REGION Network 6: GET NEXT STATION
   RUNG wire#powerrail
      P_Contact(operand := #settings.viewingStation.next.actuate, bit := #old.nextPress)
      wire#w1
      { S7_Templates := "SrcType := Int" } NE_Contact(in1 := #settings.stations.selCount, in2 := 0)
      "Get Station Selection Number"(next := TRUE, prev := FALSE, stations := #stations, selStnNumber := #settings.stations.selNumber)
   END_RUNG
   RUNG wire#powerrail
      { S7_Templates := "SrcType := Int" } NE_Contact(in1 := #settings.stations.selCount, in2 := #old.selStnCount)
   END_RUNG wire#w1
   // the same network as SCL:
   #_w1 := #settings.viewingStation.next.actuate AND NOT #old.nextPress;   // rising edge of #settings.viewingStation.next.actuate
   #old.nextPress := #settings.viewingStation.next.actuate;
   IF (#_w1 OR (#settings.stations.selCount <> #old.selStnCount)) AND (#settings.stations.selCount <> 0) THEN
       "Get Station Selection Number"(next := TRUE,
                               prev := FALSE,
                               stations := #stations,
                               selStnNumber := #settings.stations.selNumber);
   END_IF;
END_REGION

REGION Network 7: ANIMATE: NEXT STATION BUTTON
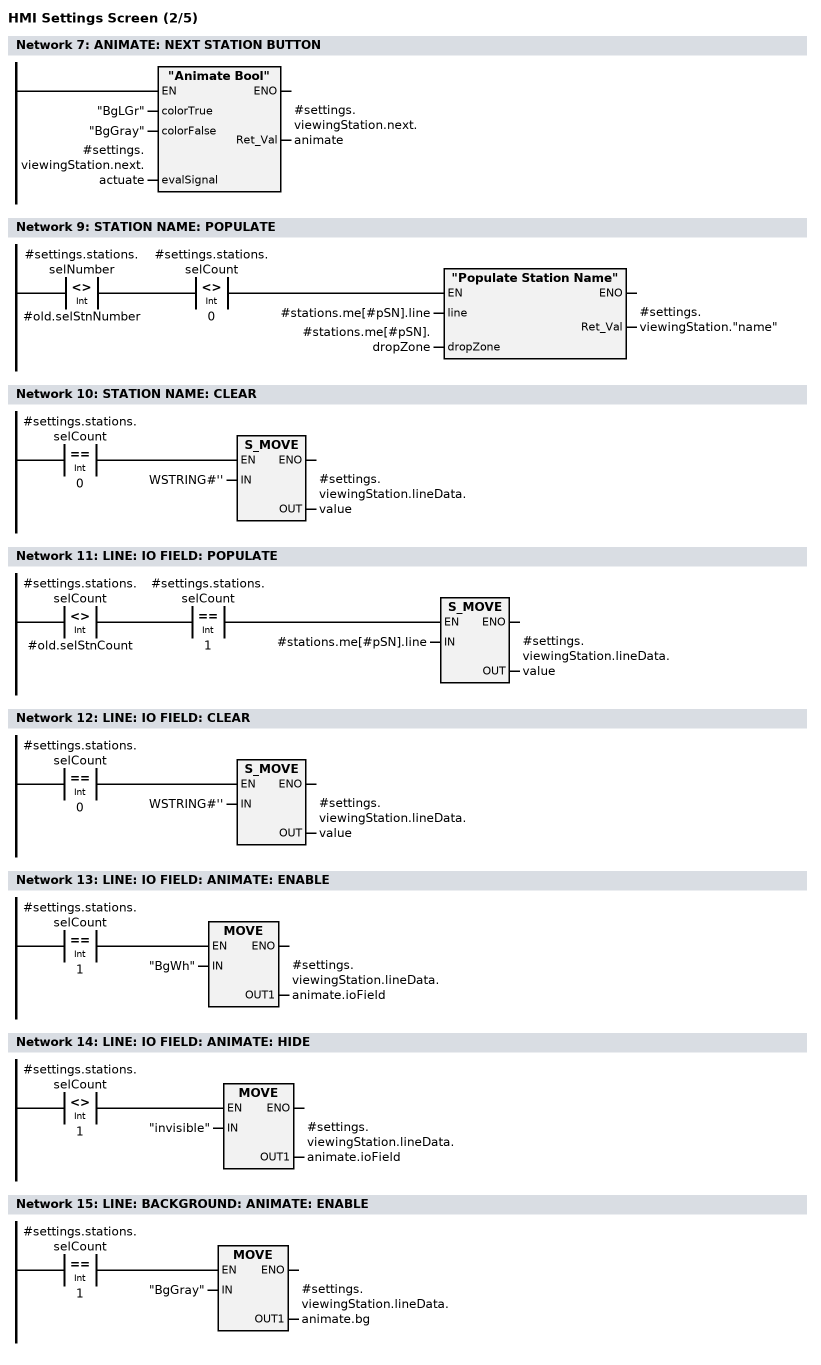
   RUNG wire#powerrail
      "Animate Bool"(colorTrue := "BgLGr", colorFalse := "BgGray", evalSignal := #settings.viewingStation.next.actuate, Ret_Val => #settings.viewingStation.next.animate)
   END_RUNG
   // the same network as SCL:
   #settings.viewingStation.next.animate := "Animate Bool"(colorTrue := "BgLGr",
                           colorFalse := "BgGray",
                           evalSignal := #settings.viewingStation.next.actuate);
END_REGION

REGION Network 8 (SCL): COPY TO POINTERS
   #pSN := #settings.stations.selNumber;
   #pBN := #settings.kp8.selBtnNumber;
END_REGION

REGION Network 9: STATION NAME: POPULATE
   RUNG wire#powerrail
      { S7_Templates := "SrcType := Int" } NE_Contact(in1 := #settings.stations.selNumber, in2 := #old.selStnNumber)
      { S7_Templates := "SrcType := Int" } NE_Contact(in1 := #settings.stations.selCount, in2 := 0)
      "Populate Station Name"(line := #stations.me[#pSN].line, dropZone := #stations.me[#pSN].dropZone, Ret_Val => #settings.viewingStation."name")
   END_RUNG
   // the same network as SCL:
   IF (#settings.stations.selNumber <> #old.selStnNumber) AND (#settings.stations.selCount <> 0) THEN
       #settings.viewingStation."name" := "Populate Station Name"(line := #stations.me[#pSN].line,
                               dropZone := #stations.me[#pSN].dropZone);
   END_IF;
END_REGION

REGION Network 10: STATION NAME: CLEAR
   RUNG wire#powerrail
      { S7_Templates := "SrcType := Int" } EQ_Contact(in1 := #settings.stations.selCount, in2 := 0)
      S_Move(in := WSTRING#'', out => #settings.viewingStation.lineData.value)
   END_RUNG
   // the same network as SCL:
   IF #settings.stations.selCount = 0 THEN #settings.viewingStation.lineData.value := WSTRING#''; END_IF;
END_REGION

REGION Network 11: LINE: IO FIELD: POPULATE
   RUNG wire#powerrail
      { S7_Templates := "SrcType := Int" } NE_Contact(in1 := #settings.stations.selCount, in2 := #old.selStnCount)
      { S7_Templates := "SrcType := Int" } EQ_Contact(in1 := #settings.stations.selCount, in2 := 1)
      S_Move(in := #stations.me[#pSN].line, out => #settings.viewingStation.lineData.value)
   END_RUNG
   // the same network as SCL:
   IF (#settings.stations.selCount <> #old.selStnCount) AND (#settings.stations.selCount = 1) THEN
       #settings.viewingStation.lineData.value := #stations.me[#pSN].line;
   END_IF;
END_REGION

REGION Network 12: LINE: IO FIELD: CLEAR
   RUNG wire#powerrail
      { S7_Templates := "SrcType := Int" } EQ_Contact(in1 := #settings.stations.selCount, in2 := 0)
      S_Move(in := WSTRING#'', out => #settings.viewingStation.lineData.value)
   END_RUNG
   // the same network as SCL:
   IF #settings.stations.selCount = 0 THEN #settings.viewingStation.lineData.value := WSTRING#''; END_IF;
END_REGION

REGION Network 13: LINE: IO FIELD: ANIMATE: ENABLE
   RUNG wire#powerrail
      { S7_Templates := "SrcType := Int" } EQ_Contact(in1 := #settings.stations.selCount, in2 := 1)
      Move(in := "BgWh", out1 => #settings.viewingStation.lineData.animate.ioField)
   END_RUNG
   // the same network as SCL:
   IF #settings.stations.selCount = 1 THEN
       #settings.viewingStation.lineData.animate.ioField := "BgWh";
   END_IF;
END_REGION

REGION Network 14: LINE: IO FIELD: ANIMATE: HIDE
   RUNG wire#powerrail
      { S7_Templates := "SrcType := Int" } NE_Contact(in1 := #settings.stations.selCount, in2 := 1)
      Move(in := "invisible", out1 => #settings.viewingStation.lineData.animate.ioField)
   END_RUNG
   // the same network as SCL:
   IF #settings.stations.selCount <> 1 THEN
       #settings.viewingStation.lineData.animate.ioField := "invisible";
   END_IF;
END_REGION

REGION Network 15: LINE: BACKGROUND: ANIMATE: ENABLE
   RUNG wire#powerrail
      { S7_Templates := "SrcType := Int" } EQ_Contact(in1 := #settings.stations.selCount, in2 := 1)
      Move(in := "BgGray", out1 => #settings.viewingStation.lineData.animate.bg)
   END_RUNG
   // the same network as SCL:
   IF #settings.stations.selCount = 1 THEN #settings.viewingStation.lineData.animate.bg := "BgGray"; END_IF;
END_REGION

REGION Network 16: LINE: BACKGROUND: ANIMATE: HIDE
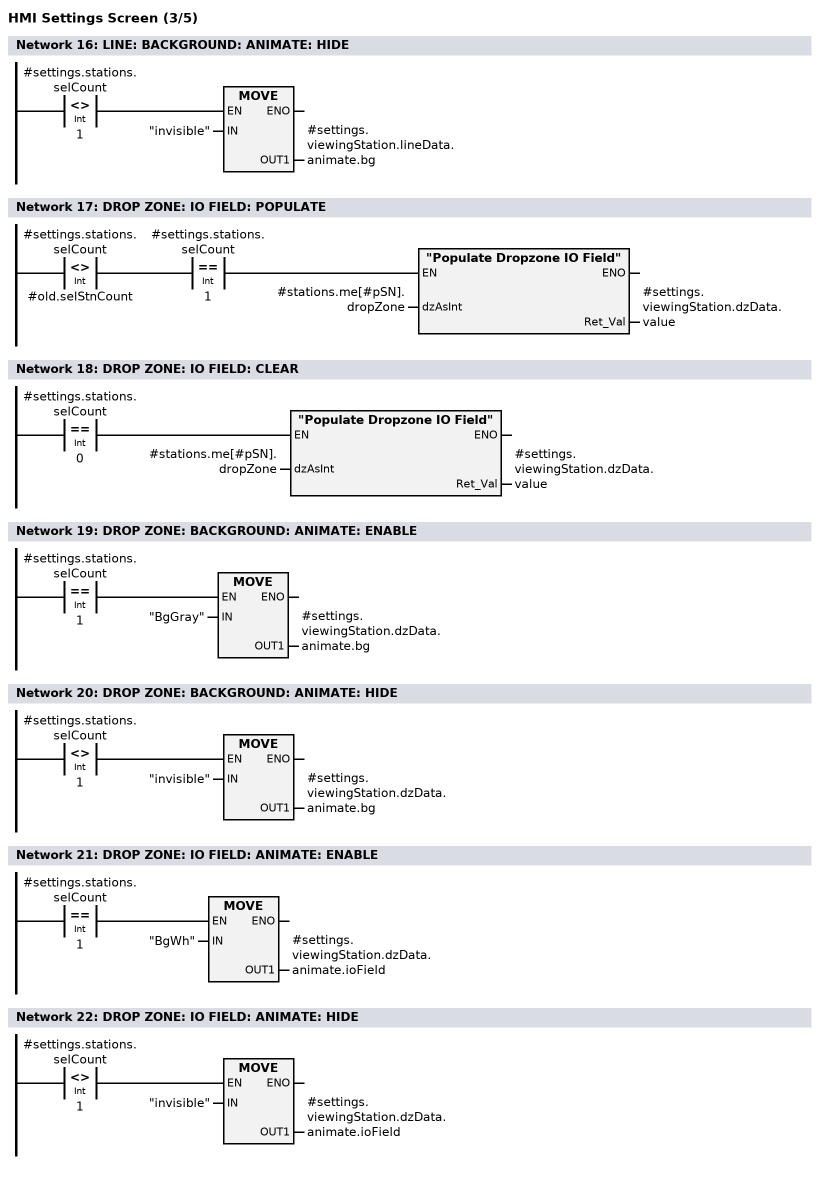
   RUNG wire#powerrail
      { S7_Templates := "SrcType := Int" } NE_Contact(in1 := #settings.stations.selCount, in2 := 1)
      Move(in := "invisible", out1 => #settings.viewingStation.lineData.animate.bg)
   END_RUNG
   // the same network as SCL:
   IF #settings.stations.selCount <> 1 THEN
       #settings.viewingStation.lineData.animate.bg := "invisible";
   END_IF;
END_REGION

REGION Network 17: DROP ZONE: IO FIELD: POPULATE
   RUNG wire#powerrail
      { S7_Templates := "SrcType := Int" } NE_Contact(in1 := #settings.stations.selCount, in2 := #old.selStnCount)
      { S7_Templates := "SrcType := Int" } EQ_Contact(in1 := #settings.stations.selCount, in2 := 1)
      "Populate Dropzone IO Field"(dzAsInt := #stations.me[#pSN].dropZone, Ret_Val => #settings.viewingStation.dzData.value)
   END_RUNG
   // the same network as SCL:
   IF (#settings.stations.selCount <> #old.selStnCount) AND (#settings.stations.selCount = 1) THEN
       #settings.viewingStation.dzData.value := "Populate Dropzone IO Field"(dzAsInt := #stations.me[#pSN].dropZone);
   END_IF;
END_REGION

REGION Network 18: DROP ZONE: IO FIELD: CLEAR
   RUNG wire#powerrail
      { S7_Templates := "SrcType := Int" } EQ_Contact(in1 := #settings.stations.selCount, in2 := 0)
      "Populate Dropzone IO Field"(dzAsInt := #stations.me[#pSN].dropZone, Ret_Val => #settings.viewingStation.dzData.value)
   END_RUNG
   // the same network as SCL:
   IF #settings.stations.selCount = 0 THEN
       #settings.viewingStation.dzData.value := "Populate Dropzone IO Field"(dzAsInt := #stations.me[#pSN].dropZone);
   END_IF;
END_REGION

REGION Network 19: DROP ZONE: BACKGROUND: ANIMATE: ENABLE
   RUNG wire#powerrail
      { S7_Templates := "SrcType := Int" } EQ_Contact(in1 := #settings.stations.selCount, in2 := 1)
      Move(in := "BgGray", out1 => #settings.viewingStation.dzData.animate.bg)
   END_RUNG
   // the same network as SCL:
   IF #settings.stations.selCount = 1 THEN #settings.viewingStation.dzData.animate.bg := "BgGray"; END_IF;
END_REGION

REGION Network 20: DROP ZONE: BACKGROUND: ANIMATE: HIDE
   RUNG wire#powerrail
      { S7_Templates := "SrcType := Int" } NE_Contact(in1 := #settings.stations.selCount, in2 := 1)
      Move(in := "invisible", out1 => #settings.viewingStation.dzData.animate.bg)
   END_RUNG
   // the same network as SCL:
   IF #settings.stations.selCount <> 1 THEN
       #settings.viewingStation.dzData.animate.bg := "invisible";
   END_IF;
END_REGION

REGION Network 21: DROP ZONE: IO FIELD: ANIMATE: ENABLE
   RUNG wire#powerrail
      { S7_Templates := "SrcType := Int" } EQ_Contact(in1 := #settings.stations.selCount, in2 := 1)
      Move(in := "BgWh", out1 => #settings.viewingStation.dzData.animate.ioField)
   END_RUNG
   // the same network as SCL:
   IF #settings.stations.selCount = 1 THEN #settings.viewingStation.dzData.animate.ioField := "BgWh"; END_IF;
END_REGION

REGION Network 22: DROP ZONE: IO FIELD: ANIMATE: HIDE
   RUNG wire#powerrail
      { S7_Templates := "SrcType := Int" } NE_Contact(in1 := #settings.stations.selCount, in2 := 1)
      Move(in := "invisible", out1 => #settings.viewingStation.dzData.animate.ioField)
   END_RUNG
   // the same network as SCL:
   IF #settings.stations.selCount <> 1 THEN
       #settings.viewingStation.dzData.animate.ioField := "invisible";
   END_IF;
END_REGION

REGION Network 23: PART NUMBER IO FIELD: POPULATE
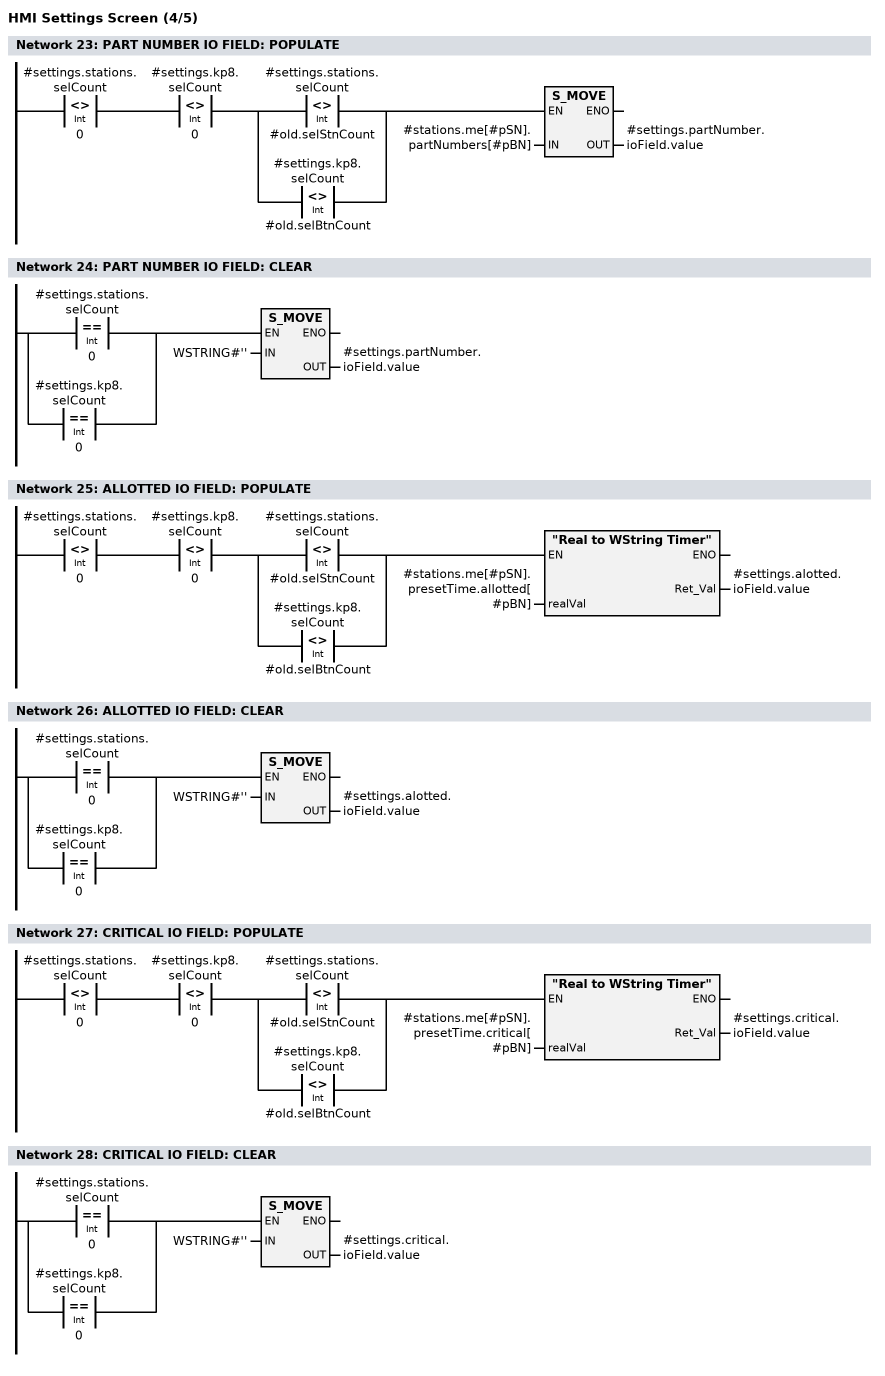
   RUNG wire#powerrail
      { S7_Templates := "SrcType := Int" } NE_Contact(in1 := #settings.stations.selCount, in2 := 0)
      { S7_Templates := "SrcType := Int" } NE_Contact(in1 := #settings.kp8.selCount, in2 := 0)
      wire#w1
      { S7_Templates := "SrcType := Int" } NE_Contact(in1 := #settings.stations.selCount, in2 := #old.selStnCount)
      wire#w2
      S_Move(in := #stations.me[#pSN].partNumbers[#pBN], out => #settings.partNumber.ioField.value)
   END_RUNG
   RUNG wire#w1
      { S7_Templates := "SrcType := Int" } NE_Contact(in1 := #settings.kp8.selCount, in2 := #old.selBtnCount)
   END_RUNG wire#w2
   // the same network as SCL:
   IF (#settings.stations.selCount <> 0) AND (#settings.kp8.selCount <> 0) AND ((#settings.stations.selCount <> #old.selStnCount) OR (#settings.kp8.selCount <> #old.selBtnCount)) THEN
       #settings.partNumber.ioField.value := #stations.me[#pSN].partNumbers[#pBN];
   END_IF;
END_REGION

REGION Network 24: PART NUMBER IO FIELD: CLEAR
   RUNG wire#powerrail
      { S7_Templates := "SrcType := Int" } EQ_Contact(in1 := #settings.stations.selCount, in2 := 0)
      wire#w1
      S_Move(in := WSTRING#'', out => #settings.partNumber.ioField.value)
   END_RUNG
   RUNG wire#powerrail
      { S7_Templates := "SrcType := Int" } EQ_Contact(in1 := #settings.kp8.selCount, in2 := 0)
   END_RUNG wire#w1
   // the same network as SCL:
   IF (#settings.stations.selCount = 0) OR (#settings.kp8.selCount = 0) THEN
       #settings.partNumber.ioField.value := WSTRING#'';
   END_IF;
END_REGION

REGION Network 25: ALLOTTED IO FIELD: POPULATE
   RUNG wire#powerrail
      { S7_Templates := "SrcType := Int" } NE_Contact(in1 := #settings.stations.selCount, in2 := 0)
      { S7_Templates := "SrcType := Int" } NE_Contact(in1 := #settings.kp8.selCount, in2 := 0)
      wire#w1
      { S7_Templates := "SrcType := Int" } NE_Contact(in1 := #settings.stations.selCount, in2 := #old.selStnCount)
      wire#w2
      "Real to WString Timer"(realVal := #stations.me[#pSN].presetTime.allotted[#pBN], Ret_Val => #settings.alotted.ioField.value)
   END_RUNG
   RUNG wire#w1
      { S7_Templates := "SrcType := Int" } NE_Contact(in1 := #settings.kp8.selCount, in2 := #old.selBtnCount)
   END_RUNG wire#w2
   // the same network as SCL:
   IF (#settings.stations.selCount <> 0) AND (#settings.kp8.selCount <> 0) AND ((#settings.stations.selCount <> #old.selStnCount) OR (#settings.kp8.selCount <> #old.selBtnCount)) THEN
       #settings.alotted.ioField.value := "Real to WString Timer"(realVal := #stations.me[#pSN].presetTime.allotted[#pBN]);
   END_IF;
END_REGION

REGION Network 26: ALLOTTED IO FIELD: CLEAR
   RUNG wire#powerrail
      { S7_Templates := "SrcType := Int" } EQ_Contact(in1 := #settings.stations.selCount, in2 := 0)
      wire#w1
      S_Move(in := WSTRING#'', out => #settings.alotted.ioField.value)
   END_RUNG
   RUNG wire#powerrail
      { S7_Templates := "SrcType := Int" } EQ_Contact(in1 := #settings.kp8.selCount, in2 := 0)
   END_RUNG wire#w1
   // the same network as SCL:
   IF (#settings.stations.selCount = 0) OR (#settings.kp8.selCount = 0) THEN
       #settings.alotted.ioField.value := WSTRING#'';
   END_IF;
END_REGION

REGION Network 27: CRITICAL IO FIELD: POPULATE
   RUNG wire#powerrail
      { S7_Templates := "SrcType := Int" } NE_Contact(in1 := #settings.stations.selCount, in2 := 0)
      { S7_Templates := "SrcType := Int" } NE_Contact(in1 := #settings.kp8.selCount, in2 := 0)
      wire#w1
      { S7_Templates := "SrcType := Int" } NE_Contact(in1 := #settings.stations.selCount, in2 := #old.selStnCount)
      wire#w2
      "Real to WString Timer"(realVal := #stations.me[#pSN].presetTime.critical[#pBN], Ret_Val => #settings.critical.ioField.value)
   END_RUNG
   RUNG wire#w1
      { S7_Templates := "SrcType := Int" } NE_Contact(in1 := #settings.kp8.selCount, in2 := #old.selBtnCount)
   END_RUNG wire#w2
   // the same network as SCL:
   IF (#settings.stations.selCount <> 0) AND (#settings.kp8.selCount <> 0) AND ((#settings.stations.selCount <> #old.selStnCount) OR (#settings.kp8.selCount <> #old.selBtnCount)) THEN
       #settings.critical.ioField.value := "Real to WString Timer"(realVal := #stations.me[#pSN].presetTime.critical[#pBN]);
   END_IF;
END_REGION

REGION Network 28: CRITICAL IO FIELD: CLEAR
   RUNG wire#powerrail
      { S7_Templates := "SrcType := Int" } EQ_Contact(in1 := #settings.stations.selCount, in2 := 0)
      wire#w1
      S_Move(in := WSTRING#'', out => #settings.critical.ioField.value)
   END_RUNG
   RUNG wire#powerrail
      { S7_Templates := "SrcType := Int" } EQ_Contact(in1 := #settings.kp8.selCount, in2 := 0)
   END_RUNG wire#w1
   // the same network as SCL:
   IF (#settings.stations.selCount = 0) OR (#settings.kp8.selCount = 0) THEN
       #settings.critical.ioField.value := WSTRING#'';
   END_IF;
END_REGION

REGION Network 29: PART NUMBER, ALLOTTED & CRITICAL: ANIMATE
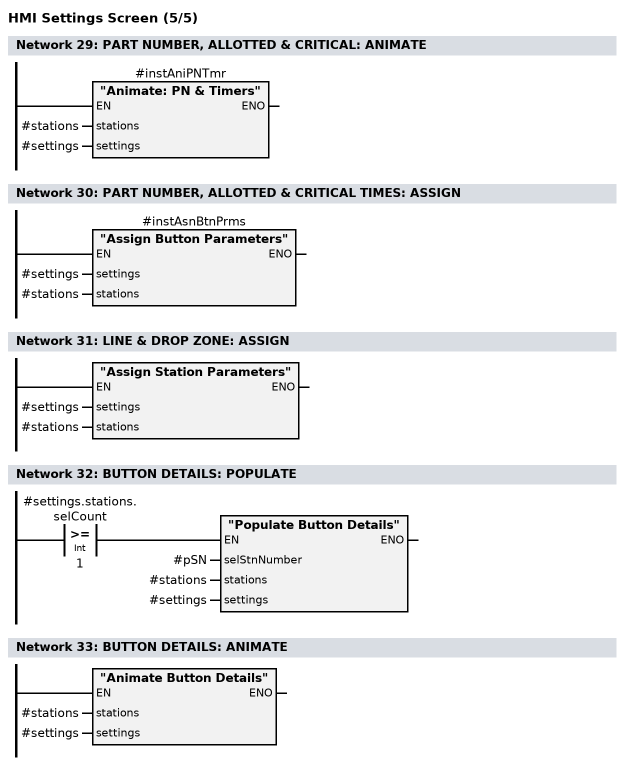
   RUNG wire#powerrail
      #instAniPNTmr(stations := #stations, settings := #settings)
   END_RUNG
   // the same network as SCL:
   #instAniPNTmr(stations := #stations, settings := #settings);   // "Animate: PN & Timers"
END_REGION

REGION Network 30: PART NUMBER, ALLOTTED & CRITICAL TIMES: ASSIGN
   RUNG wire#powerrail
      #instAsnBtnPrms(settings := #settings, stations := #stations)
   END_RUNG
   // the same network as SCL:
   #instAsnBtnPrms(settings := #settings, stations := #stations);   // "Assign Button Parameters"
END_REGION

REGION Network 31: LINE & DROP ZONE: ASSIGN
   RUNG wire#powerrail
      "Assign Station Parameters"(settings := #settings, stations := #stations)
   END_RUNG
   // the same network as SCL:
   "Assign Station Parameters"(settings := #settings, stations := #stations);
END_REGION

REGION Network 32: BUTTON DETAILS: POPULATE
   RUNG wire#powerrail
      { S7_Templates := "SrcType := Int" } GE_Contact(in1 := #settings.stations.selCount, in2 := 1)
      "Populate Button Details"(selStnNumber := #pSN, stations := #stations, settings := #settings)
   END_RUNG
   // the same network as SCL:
   IF #settings.stations.selCount >= 1 THEN
       "Populate Button Details"(selStnNumber := #pSN, stations := #stations, settings := #settings);
   END_IF;
END_REGION

REGION Network 33: BUTTON DETAILS: ANIMATE
   RUNG wire#powerrail
      "Animate Button Details"(stations := #stations, settings := #settings)
   END_RUNG
   // the same network as SCL:
   "Animate Button Details"(stations := #stations, settings := #settings);
END_REGION

REGION Network 34 (SCL): CHANGE DETECTION
   #old.selBtnCount := #settings.kp8.selCount;
   #old.selBtnNumber := #settings.kp8.selBtnNumber;
   #old.selStnCount := #settings.stations.selCount;
   #old.selStnNumber := #settings.stations.selNumber;
END_REGION
END_FUNCTION_BLOCK

FUNCTION_BLOCK "HMI Populate Part Call"   // FB16, SCL
{ S7_Optimized_Access := 'TRUE' }
VERSION : 0.1
   VAR_INPUT
      firstScan : Bool;
      currentRowCount : Int;
      requests : "Part Request Data";
   END_VAR
   VAR_IN_OUT
      partCall : "Part Call Screen";
      tableNav : "Table Nav";
   END_VAR
   VAR
      firstRow : Int;
      old : Struct
         top : Bool;
         pgUp : Bool;
         lnUp : Bool;
         lnDn : Bool;
         pgDn : Bool;
         btm : Bool;
      END_STRUCT;
   END_VAR
   VAR_TEMP
      animate : Bool;
      btn : Struct
         top : Bool;
         pgUp : Bool;
         lnUp : Bool;
         lnDn : Bool;
         pgDn : Bool;
         btm : Bool;
      END_STRUCT;
      gray : USInt;
      green : USInt;
      i : Int;
      maxDBRows : Int;
      pRow : Int;
      visibleRows : Int;
      thisRow : Int;
      saveAct : Bool;
   END_VAR
BEGIN
   REGION "COPY TO LOCAL"
       #visibleRows := "partReqHmiRowCount";
       #maxDBRows := #currentRowCount;
       #btn.top := #tableNav.top.actuate;
       #btn.pgUp := #tableNav.pageUp.actuate;
       #btn.lnUp := #tableNav.lineUp.actuate;
       #btn.lnDn := #tableNav.lineDown.actuate;
       #btn.pgDn := #tableNav.pageDown.actuate;
       #btn.btm := #tableNav.bottom.actuate;
   END_REGION

   REGION "RESOLVE FIRST ROW"

       REGION "TOP"
           IF NOT #btn.top AND #old.top THEN
               #firstRow := 0;
           END_IF;
       END_REGION

       REGION "PAGE UP"
           IF NOT #btn.pgUp AND #old.pgUp THEN
               #firstRow -= #visibleRows - 1;
           END_IF;
       END_REGION

       REGION "LINE UP"
           IF NOT #btn.lnUp AND #old.lnUp THEN
               #firstRow -= 1;
           END_IF;
       END_REGION

       REGION "LINE DOWN"
           IF NOT #btn.lnDn AND #old.lnDn THEN
               #firstRow += 1;
           END_IF;
       END_REGION

       REGION "PAGE DOWN"
           IF NOT #btn.pgDn AND #old.pgDn THEN
               #firstRow += #visibleRows - 1;
           END_IF;
       END_REGION

       REGION "BOTTOM"
           IF NOT #btn.btm AND #old.btm THEN
               #firstRow := #maxDBRows - #visibleRows + 1;
           END_IF;
       END_REGION

   END_REGION

   REGION "CHANGE DETECTION"
       #old.top := #btn.top;
       #old.pgUp := #btn.pgUp;
       #old.lnUp := #btn.lnUp;
       #old.lnDn := #btn.lnDn;
       #old.pgDn := #btn.pgDn;
       #old.btm := #btn.btm;
   END_REGION

   REGION "ANIMATE PART CALL NAV"

       REGION "COPY TO LOCAL"
           #gray := "BgGray";
           #green := "BgLGr";
       END_REGION

       REGION "TOP"
           #tableNav.top.animate := "Animate Bool"(colorTrue := #green,
                                                   colorFalse := #gray,
                                                   evalSignal := #tableNav.top.actuate);
       END_REGION

       REGION "PAGE UP"
           #tableNav.pageUp.animate := "Animate Bool"(colorTrue := #green,
                                                      colorFalse := #gray,
                                                      evalSignal := #tableNav.pageUp.actuate);
       END_REGION

       REGION "LINE UP"
           #tableNav.lineUp.animate := "Animate Bool"(colorTrue := #green,
                                                      colorFalse := #gray,
                                                      evalSignal := #tableNav.lineUp.actuate);
       END_REGION

       REGION "LINE DOWN"
           #tableNav.lineDown.animate := "Animate Bool"(colorTrue := #green,
                                                        colorFalse := #gray,
                                                        evalSignal := #tableNav.lineDown.actuate);
       END_REGION

       REGION "PAGE DOWN"
           #tableNav.pageDown.animate := "Animate Bool"(colorTrue := #green,
                                                        colorFalse := #gray,
                                                        evalSignal := #tableNav.pageDown.actuate);
       END_REGION

       REGION "BOTTOM"
           #tableNav.bottom.animate := "Animate Bool"(colorTrue := #green,
                                                      colorFalse := #gray,
                                                      evalSignal := #tableNav.bottom.actuate);
       END_REGION

   END_REGION

   REGION "UPPER LIMIT ROLL OVER"
       IF #firstRow > #maxDBRows THEN
           #firstRow -= #maxDBRows - 1;
       END_IF;
   END_REGION

   REGION "LOWER LIMIT ROLL OVER"
       IF #firstRow < 0 THEN
           #firstRow += #maxDBRows - 1;
       END_IF;
   END_REGION

   REGION "LOOP THROUGH DISPLAYED STATIONS"
       FOR #i := 0 TO #visibleRows - 1 DO

           REGION "CALCULATE POINTER"
               #pRow := #firstRow + #i;
           END_REGION

           REGION "UPPER LIMIT ROLL OVER"
               IF #maxDBRows <= #visibleRows THEN
                   #pRow := #i;
               END_IF;
               IF #pRow >= #maxDBRows AND #maxDBRows >= #visibleRows THEN
                   #pRow := #firstRow + #i - #maxDBRows;
               END_IF;
           END_REGION

           REGION "SEND TO HMI"
               #saveAct := #partCall.row[#i].pbSelection.actuate;
               #partCall.row[#i] := #requests.row[#pRow];
               #partCall.row[#i].pbSelection.actuate := #saveAct;
           END_REGION

       END_FOR;
   END_REGION
END_FUNCTION_BLOCK

FUNCTION_BLOCK "Load Default Timer Presets"   // FB18, SCL
{ S7_Optimized_Access := 'TRUE' }
VERSION : 0.1
   VAR_INPUT
      req : Bool;
   END_VAR
   VAR_IN_OUT
      stations : "Stations";
   END_VAR
   VAR
      oldReq : Bool;
   END_VAR
   VAR_TEMP
      alotted : Real;
      critical : Real;
      i : Int;
      j : Int;
      partNumber : WString;
      tmrReal : Real;
   END_VAR
BEGIN
   REGION "COPY TO LOCAL"
       #alotted := "defaultAlotted";
       #critical := "defaultCritical";
   END_REGION

   REGION "ON REQUEST RISING EDGE"
       IF #req AND NOT #oldReq THEN

           REGION "LOOP THROUGH STATIONS" 
               FOR #i := 0 TO "stnCount" DO

                   REGION "LOOP THROUGH BUTTONS"
                       FOR #j := 0 TO "ptsPerStn" DO

                           REGION "COPY TO LOCAL"
                               #partNumber := #stations.me[#i].partNumbers[#j];
                           END_REGION

                           REGION "IF BUTTON HAS ASSOCIATED PN"
                               IF LEN(#partNumber) <> 0 THEN

                                   REGION "COPY TO LOCAL"
                                       #tmrReal := #stations.me[#i].presetTime.allotted[#j];
                                   END_REGION

                                   REGION "ON NO TIME ENTERED"
                                       IF #tmrReal = 0.0 THEN

                                           REGION "ASSIGN ALLOTTED VALUES"
                                               #stations.me[#i].presetTime.allotted[#j] := #alotted;
                                           END_REGION

                                       END_IF;
                                   END_REGION

                                   REGION "COPY TO LOCAL"
                                       #tmrReal := #stations.me[#i].presetTime.critical[#j];
                                   END_REGION

                                   REGION "ON NO TIME ENTERED"
                                       IF #tmrReal = 0.0 THEN

                                           REGION "ASSIGN CRITICAL VALUES"
                                               #stations.me[#i].presetTime.critical[#j] := #critical;
                                           END_REGION

                                       END_IF;
                                   END_REGION

                               END_IF;
                           END_REGION

                       END_FOR;
                   END_REGION

               END_FOR;
           END_REGION

       END_IF;
   END_REGION

   REGION "CHANGE DETECTION"
       #oldReq := #req;
   END_REGION ;
END_FUNCTION_BLOCK

FUNCTION_BLOCK "LED Populate Sign"   // FB19, SCL
{ S7_Optimized_Access := 'TRUE' }
VERSION : 0.1
   VAR_INPUT
      requests : "Part Request Data";
   END_VAR
   VAR_IN_OUT
      ledData : "LED Sign Data";
   END_VAR
   VAR_TEMP
      animate : USInt;
      i : Int;
      visibleRows : Int;
      tempRow : "Table Row";
   END_VAR
BEGIN
   REGION "COPY TO LOCAL"
       #visibleRows := "ledRowCount";
   END_REGION

   REGION "POPULATE SIGN DATA"

       REGION "FOR EACH ROW ON SIGN"
           FOR #i := 0 TO #visibleRows DO

               REGION "GET ROW"
                   #tempRow := #requests.row[#i];
               END_REGION

               REGION "LINE LABEL DARK MODE"                
                   "Dark Mode"(#tempRow.tfLine.animate);
               END_REGION

               REGION "DROP ZONE DARK MODE"
                   "Dark Mode"(#tempRow.tfDropZone.animate);
               END_REGION

               REGION "PART NUMBER DARK MODE"

                   REGION "SINGLE LINE"
                       "Dark Mode"(#tempRow.tfPartNumber.animateSL);
                   END_REGION

                   REGION "DOUBLE LINE"
                       "Dark Mode"(#tempRow.tfPartNumber.animateDL);
                   END_REGION

               END_REGION

               REGION "TIME DARK MODE"
                   "Dark Mode"(#tempRow.tfTime.animate);
               END_REGION

               REGION "SEND TO SIGN"
                   #ledData.row[#i] := #tempRow;
               END_REGION

           END_FOR;
       END_REGION

   END_REGION
END_FUNCTION_BLOCK

FUNCTION_BLOCK "Station Selection"   // FB20, SCL
{ S7_Optimized_Access := 'TRUE' }
VERSION : 0.1
   VAR_IN_OUT
      settings : "Settings";
      stations : "Stations";
   END_VAR
   VAR
      firstStn : Int;
      rt : "Runtime Data";
      selectionExe : Bool;
      old : Struct
         prevGrp : Bool;
         nextGrp : Bool;
         stnSlct : Array[0..11] of Bool;
      END_STRUCT;
   END_VAR
   VAR_TEMP
      animate : USInt;
      btnPress : Bool;
      count : Int;
      currentBtn : Bool;
      evalObjCount : Int;
      i : Int;
      oldBtn : Bool;
      pStn : Int;
      stnName : WString;
      stnSelected : Bool;
      selState : Bool;
      selStnCount : Int;
      timerExpired : Bool;
      stnSelLblCount : Int;
   END_VAR
   VAR CONSTANT
      ptTimer : Real := 1.5;
   END_VAR
BEGIN
   REGION "UI INTERACTION ANIMATIONS"

       REGION "NEXT GROUP"
           #btnPress := #settings.stations.nextGroup.actuate;
           #animate := "Animate Bool"(colorTrue := "BgLGr",
                                      colorFalse := "BgGray",
                                      evalSignal := #btnPress);
           #settings.stations.nextGroup.animate := #animate;
       END_REGION

       REGION "PREVIOUS GROUP"
           #btnPress := #settings.stations.prevGroup.actuate;
           #animate := "Animate Bool"(colorTrue := "BgLGr",
                                      colorFalse := "BgGray",
                                      evalSignal := #btnPress);
           #settings.stations.prevGroup.animate := #animate;
       END_REGION

       REGION "SELECT ALL STATIONS"
           #btnPress := #settings.stations.selectAll.actuate;
           #animate := "Animate Bool"(colorTrue := "BgLGr",
                                      colorFalse := "BgGray",
                                      evalSignal := #settings.stations.selectAll.actuate);
           #settings.stations.selectAll.animate := #animate;
       END_REGION

   END_REGION

   REGION "POPULATE STATION LABELS"

       REGION "PROCESS NEXT GROUP PRESS"

           REGION "COPY TO LOCAL"
               #currentBtn := #settings.stations.nextGroup.actuate;
               #oldBtn := #old.nextGrp;
           END_REGION

           REGION "FALLING EDGE OF NEXT GROUP"
               IF NOT #currentBtn AND #oldBtn THEN

                   REGION "INCREMENT FIRST STATION"
                       #firstStn := #firstStn + 2;
                   END_REGION

                   REGION "UPPER LIMIT ROLL OVER"
                       IF #firstStn > "stnCount" THEN
                           #firstStn := #firstStn - "stnCount" - 1;
                       END_IF;
                   END_REGION

               END_IF;
           END_REGION

           REGION "NEXT GROUP CHANGE DETECTION"
               #old.nextGrp := #currentBtn;
           END_REGION

       END_REGION

       REGION "PROCESS PREVIOUS GROUP PRESS"

           REGION "COPY TO LOCAL"
               #currentBtn := #settings.stations.prevGroup.actuate;
               #oldBtn := #old.prevGrp;
           END_REGION

           REGION "FALLING EDGE OF PREVIOUS GROUP"
               IF NOT #currentBtn AND #oldBtn THEN

                   REGION "DECREMENT FIRST STATION"
                       #firstStn := #firstStn - 2;
                   END_REGION

                   REGION "LOWER LIMIT ROLL OVER"
                       IF #firstStn < 0 THEN
                           #firstStn := #firstStn + "stnCount" + 1;
                       END_IF;
                   END_REGION

               END_IF;
           END_REGION

           REGION "PREVIOUS GROUP CHANGE DETECTION"
               #old.prevGrp := #currentBtn;
           END_REGION

       END_REGION

       REGION "WRITE LABEL"

           REGION "COPY TO LOCAL"
               #evalObjCount := "hmiSelStnCount";
           END_REGION

           REGION "FOR EACH STATION SELECTION BUTTON"
               FOR #i := 0 TO #evalObjCount DO

                   REGION "CALCULATE POINTER"
                       #pStn := #firstStn + #i;
                   END_REGION

                   REGION "UPPER LIMIT ROLL OVER"
                       IF #pStn > "stnCount" THEN
                           #pStn := #firstStn + #i - "stnCount" - 1;
                       END_IF;
                   END_REGION

                   REGION "BUILD NAME"
                       #stnName := CONCAT_WSTRING(IN1 := #stations.me[#pStn].line,
                                                  IN2 := wstring#' ',
                                                  IN3 := "Strip Sign"(USINT_TO_WSTRING(#stations.me[#pStn].dropZone)));
                   END_REGION

                   REGION "WRITE NAME"
                       #settings.stations.selectBtns[#i].label := #stnName;
                   END_REGION

               END_FOR;
           END_REGION

       END_REGION

   END_REGION

   REGION "SINGLE STATION SELECTION"

       REGION "COPY TO LOCAL"
           #stnSelLblCount := "hmiSelStnCount";
       END_REGION

       REGION "LOOP THROUGH DISPLAYED STATIONS"
           FOR #i := 0 TO #stnSelLblCount DO

               REGION "CALCULATE POINTER"
                   #pStn := #firstStn + #i;
               END_REGION

               REGION "UPPER LIMIT ROLL OVER"
                   IF #pStn > "stnCount" THEN
                       #pStn := #firstStn + #i - "stnCount" - 1;
                   END_IF;
               END_REGION

               REGION "COPY TO LOCAL"
                   #currentBtn := #settings.stations.selectBtns[#i].actuate;
                   #oldBtn := #old.stnSlct[#i];
               END_REGION

               REGION "TOGGLE STATE ON FALLING EDGE"
                   IF NOT #currentBtn AND #oldBtn THEN
                       #selState := #stations.me[#pStn].settings.selected;
                       #selState := NOT #selState;
                       #stations.me[#pStn].settings.selected := #selState;
                   END_IF;
               END_REGION

               REGION "STATION SELECTION CHANGE DETECTION"
                   #old.stnSlct[#i] := #currentBtn;
               END_REGION

           END_FOR;
       END_REGION

   END_REGION

   REGION "MULTI SELECT TIMER"

       REGION "RUNTIME CALL"
           #rt.elapsed := RUNTIME(#rt.mem);
       END_REGION

       REGION "TIMER"

           REGION "COPY TO LOCAL"
               #btnPress := #settings.stations.selectAll.actuate;
           END_REGION

           REGION "ACCUMULATE RT VALUES"
               IF #btnPress THEN
                   #rt.asReal += LREAL_TO_REAL(#rt.elapsed);
               END_IF;
           END_REGION

           REGION "SET TIMER FLAG"
               IF #rt.asReal < #ptTimer THEN
                   #timerExpired := FALSE;
               END_IF;
               IF #rt.asReal >= #ptTimer THEN
                   #timerExpired := TRUE;
                   #rt.asReal := 0.0;
               END_IF;
           END_REGION

           REGION "RESET ACCUMULATED VALUE"
               IF NOT #btnPress THEN
                   #rt.asReal := 0.0;
                   #selectionExe := FALSE;
               END_IF;
           END_REGION

       END_REGION

   END_REGION

   REGION "EVALUATE MULTI SELECTION"
       IF #timerExpired AND NOT #selectionExe THEN

           REGION "COPY TO LOCAL"
               #selStnCount := #settings.stations.selCount;
           END_REGION

           REGION "SELECT ALL"
               IF #selStnCount < "stnCount" THEN
                   "Select Stations"(mode := TRUE,
                                     stations := #stations);
               END_IF;
           END_REGION

           REGION "DESELECT ALL"
               IF #selStnCount = "stnCount" THEN
                   "Select Stations"(mode := FALSE,
                                     stations := #stations);
               END_IF;
           END_REGION

           REGION "FLAG SELECTION EXECUTED"
               #selectionExe := TRUE;
           END_REGION

       END_IF;
   END_REGION

   REGION "SELECTION ANIMATIONS"

       REGION "COPY TO LOCAL"
           #stnSelLblCount := "hmiSelStnCount";
       END_REGION

       REGION "LOOP THROUGH BUTTONS"
           FOR #i := 0 TO #stnSelLblCount DO

               REGION "CALCULATE POINTER"
                   #pStn := #firstStn + #i;
               END_REGION

               REGION "UPPER LIMIT ROLL OVER"
                   IF #pStn > "stnCount" THEN
                       #pStn := #firstStn + #i - "stnCount" - 1;
                   END_IF;
               END_REGION

               REGION "COPY TO LOCAL"
                   #currentBtn := #settings.stations.selectBtns[#i].actuate;
                   #stnSelected := #stations.me[#pStn].settings.selected;
               END_REGION

               REGION "DRAW SELCTION HIGHLIGHTS"
                   #animate := "Animate Bool"(colorTrue := "BgLTe",
                                              colorFalse := "BgGray",
                                              evalSignal := #stnSelected);
               END_REGION

               REGION "ANIMATE BUTTON PRESS"
                   #animate := "Animate Bool"(colorTrue := "BgDTe",
                                              colorFalse := #animate,
                                              evalSignal := #currentBtn);
                   #settings.stations.selectBtns[#i].animate := #animate;
               END_REGION

           END_FOR;
       END_REGION

   END_REGION

   REGION "COUNT SELECTED STATIONS"

       REGION "INITIALIZE LOCAL"
           #count := 0;
           #evalObjCount := "stnCount";
       END_REGION

       REGION "LOOP THROUGH STATIONS"
           FOR #i := 0 TO #evalObjCount DO

               REGION "INCREMENT COUNT ON SELECTION"
                   #stnSelected := #stations.me[#i].settings.selected;
                   IF #stnSelected THEN
                       #count += 1;
                   END_IF;
               END_REGION

           END_FOR;
       END_REGION

       REGION "SAVE COUNT"
           #settings.stations.selCount := #count;
       END_REGION

   END_REGION
END_FUNCTION_BLOCK

FUNCTION_BLOCK "KP8 Button Selections"   // FB21, SCL
{ S7_Optimized_Access := 'TRUE' }
VERSION : 0.1
   VAR_INPUT
      reset : Bool;
   END_VAR
   VAR_IN_OUT
      settings : "Settings";
      stations : "Stations";
   END_VAR
   VAR
      enableState : Bool;
      oldBtnPresses : Array[0..7] of Bool;
      oldSelState : Array[0..7] of Bool;
      oldSelStnCount : Int;
      rt : "Runtime Data";
      timerExpired : Bool;
      selectionExe : Bool;
   END_VAR
   VAR_TEMP
      animate : USInt;
      btnPress : Bool;
      count : Int;
      i : Int;
      j : Int;
      mode : Bool;
      oldPress : Bool;
      pBtn : Int;
      selBtnCount : Int;
      selStnCount : Int;
      stnSelected : Bool;
   END_VAR
   VAR CONSTANT
      selectAllTime : Real := 1.5;
   END_VAR
BEGIN
   REGION "ENABLE KP8 BUTTON ASSIGNMENT SECTION"

       REGION "ENABLE"

           REGION "COPY TO LOCAL"
               #selStnCount := #settings.stations.selCount;
           END_REGION

           REGION "ON CHANGE IN SELECTED STATION COUNT"
               IF #selStnCount <> 0 AND #selStnCount <> #oldSelStnCount THEN

                   REGION "ENABLE KP8 SELECTIONS"
                       #enableState := TRUE;
                   END_REGION

               END_IF;
           END_REGION

       END_REGION

       REGION "DISABLE"

           REGION "COPY TO LOCAL"
               #selStnCount := #settings.stations.selCount;
           END_REGION

           REGION "ON DESELETION OF LAST STATION"
               IF #selStnCount = 0 AND #selStnCount <> #oldSelStnCount THEN

                   REGION "RESET ENABLED STATE"
                       #enableState := FALSE;
                   END_REGION

                   REGION "RESET BUTTON SELECTION STATES"
                       FOR #i := 0 TO "ptsPerStn" DO
                           #settings.kp8.btnSelState[#i] := FALSE;
                       END_FOR;
                   END_REGION

               END_IF;
           END_REGION

       END_REGION

   END_REGION

   REGION "SINGLE BUTTON SELECTION"

       REGION "LOOP THROUGH BUTTONS"
           FOR #i := 0 TO "ptsPerStn" DO

               REGION "EXCLUDE STOP RUNTIME AND RESET SELECTED BUTTONS"
                   IF #i <> 0 AND #i <> 4 THEN

                       REGION "COPY TO LOCAL"

                           REGION "CALCULATE BUTTON POINTER"
                               CASE #i OF
                                   1:
                                       #pBtn := 5;
                                   2:
                                       #pBtn := 3;
                                   3:
                                       #pBtn := 1;
                                   5:
                                       #pBtn := 4;
                                   6:
                                       #pBtn := 2;
                                   7:
                                       #pBtn := 0;
                                   ELSE
                                       ;
                               END_CASE;
                           END_REGION

                           #btnPress := #settings.kp8.buttons[#i].actuate OR #settings.viewingStation.btns[#pBtn].select.actuate;
                           #oldPress := #oldBtnPresses[#i];

                       END_REGION

                       REGION "TOGGLE STATE ON FALLING EDGE"
                           IF NOT #btnPress AND #oldPress THEN
                               #settings.kp8.btnSelState[#i] := NOT #settings.kp8.btnSelState[#i];
                               #settings.kp8.selBtnNumber := #i;
                           END_IF;
                       END_REGION

                       REGION "SAVE SELECTED BUTTON NUMBER ON DESELECT"
                           IF NOT #settings.kp8.btnSelState[#i] AND #oldSelState[#i] THEN
                               FOR #j := 0 TO "ptsPerStn" DO
                                   IF #settings.kp8.btnSelState[#j] THEN
                                       #settings.kp8.selBtnNumber := #j;
                                   END_IF;
                               END_FOR;
                           END_IF;
                       END_REGION

                       REGION "KP8 BUTON SELECTION CHANGE DETECTION"
                           #oldBtnPresses[#i] := #btnPress;
                       END_REGION

                   END_IF;
               END_REGION

           END_FOR;
       END_REGION

   END_REGION

   REGION "MULTI BUTTON SELECTION"

       REGION "MULTI SELECT TIMER"

           REGION "RUNTIME CALL"
               #rt.elapsed := RUNTIME(#rt.mem);
           END_REGION

           REGION "TIMER"

               REGION "COPY TO LOCAL"
                   #btnPress := #settings.kp8.selectButtons.actuate;
               END_REGION

               REGION "ACCUMULATE RT VALUES"
                   IF #btnPress THEN
                       #rt.asReal += LREAL_TO_REAL(#rt.elapsed);
                   END_IF;
               END_REGION

               REGION "SET TIMER FLAG"
                   IF #rt.asReal < #selectAllTime THEN
                       #timerExpired := FALSE;
                   END_IF;
                   IF #rt.asReal >= #selectAllTime THEN
                       #timerExpired := TRUE;
                       #rt.asReal := 0.0;
                   END_IF;
               END_REGION

               REGION "RESET ACCUMULATED VALUE"
                   IF NOT #btnPress THEN
                       #rt.asReal := 0.0;
                       #selectionExe := FALSE;
                   END_IF;
               END_REGION

           END_REGION

       END_REGION

       REGION "EVALUATE MULTI SELECTION"
           IF #timerExpired AND NOT #selectionExe THEN

               REGION "COPY TO LOCAL"
                   #selBtnCount := #settings.kp8.selCount;
               END_REGION

               REGION "SELECT ALL"
                   IF #selBtnCount < "ptsPerStn" - 1 THEN
                       #mode := TRUE;
                   END_IF;
               END_REGION

               REGION "DESELECT ALL"
                   IF #selBtnCount = "ptsPerStn" - 1 THEN
                       #mode := FALSE;
                   END_IF;
               END_REGION

               REGION "SAVE SELECTIONS"
                   FOR #i := 0 TO "ptsPerStn" DO

                       REGION "EXCLUDE STOP RUNTIME AND RESET SELECTED BUTTONS"
                           IF #i <> 0 AND #i <> 4 THEN

                               REGION "PERFROM SELECTION"
                                   #settings.kp8.btnSelState[#i] := #mode;
                               END_REGION

                           END_IF;
                       END_REGION

                   END_FOR;
               END_REGION

               REGION "SET SELECED BUTTON NUMBER TO 1"
                   #settings.kp8.selBtnNumber := 0;
               END_REGION

               REGION "FLAG SELECTION EXECUTED"
                   #selectionExe := TRUE;
               END_REGION

           END_IF;
       END_REGION
   END_REGION

   REGION "SAVE BUTTON SELECTIONS TO STATIONS"

       REGION "COPY TO LOCAL"
           #selStnCount := #settings.stations.selCount;
       END_REGION

       REGION "ON CHANGE IN BUTTON OR STATION SELECTON"
           IF #settings.kp8.btnSelState <> #oldSelState OR #selStnCount <> #oldSelStnCount THEN

               REGION "FOR SELECTED STATIONS"
                   FOR #i := 0 TO "stnCount" DO
                       #stnSelected := #stations.me[#i].settings.selected;
                       IF #stnSelected THEN

                           REGION "SAVE BUTTON SELECTION STATE"
                               #stations.me[#i].settings.btnSelection := #settings.kp8.btnSelState;
                           END_REGION

                       END_IF;
                   END_FOR;
               END_REGION

           END_IF;
       END_REGION

       REGION "SELECTED STATION COUNT CHANGE DETECTION"
           #oldSelStnCount := #selStnCount; 
       END_REGION

   END_REGION

   REGION "COUNT SELECTED BUTTONS"

       REGION "ON CHANGE IN BUTTON SELECTION STATES"
           IF #settings.kp8.btnSelState <> #oldSelState THEN

               REGION "INITIALIZE LOCAL"
                   #count := 0;
               END_REGION

               REGION "FOR EACH SELECTED BUTTON"
                   FOR #i := 0 TO "ptsPerStn" DO
                       IF #settings.kp8.btnSelState[#i] THEN

                           REGION "INCREMENT COUNT"
                               #count := #count + 1;
                           END_REGION

                       END_IF;
                   END_FOR;
               END_REGION

               REGION "SAVE COUNT"
                   #settings.kp8.selCount := #count;
               END_REGION

           END_IF;
       END_REGION

   END_REGION 

   REGION "UI INTERACTION ANIMATIONS"

       REGION "SELECT ALL BUTTONS"
           #btnPress := #settings.kp8.selectButtons.actuate;
           #animate := "Animate Bool"(colorTrue := "BgLGr",
                                      colorFalse := "BgGray",
                                      evalSignal := #btnPress);
           #settings.kp8.selectButtons.animate := #animate;
       END_REGION

       REGION "STOP RESET SELECTED STATION"
           #btnPress := #settings.kp8.buttons[0].actuate;
           #animate := "Animate Bool"(colorTrue := "FgGray",
                                      colorFalse := "BgGray",
                                      evalSignal := #btnPress);
           #settings.kp8.buttons[0].animate := #animate;
       END_REGION

       REGION "STOP RUNTIME"
           #btnPress := #settings.kp8.buttons[4].actuate;
           #animate := "Animate Bool"(colorTrue := "FgGray",
                                      colorFalse := "BgGray",
                                      evalSignal := #btnPress);
           #settings.kp8.buttons[4].animate := #animate;
       END_REGION

       REGION "BUTTON SELECTIONS"

           REGION "FOR EACH BUTTON"     
               FOR #i := 0 TO "ptsPerStn" DO

                   REGION "EXCLUDE STOP RUNTIME AND RESET SELECTED BUTTONS"
                       IF #i <> 0 AND #i <> 4 THEN

                           REGION "ANIMATE"

                               REGION "COPY TO LOCAL"
                                   #btnPress := #settings.kp8.buttons[#i].actuate;
                               END_REGION

                               REGION "ENABLE/DISABLE"
                                   #animate := "Animate Bool"(colorTrue := "BgGray",
                                                              colorFalse := "disabled",
                                                              evalSignal := #enableState);
                               END_REGION

                               REGION "ENABLED SUB ANIMATIONS"
                                   IF #enableState THEN

